REGION Network 19: EM - Execute State Complete
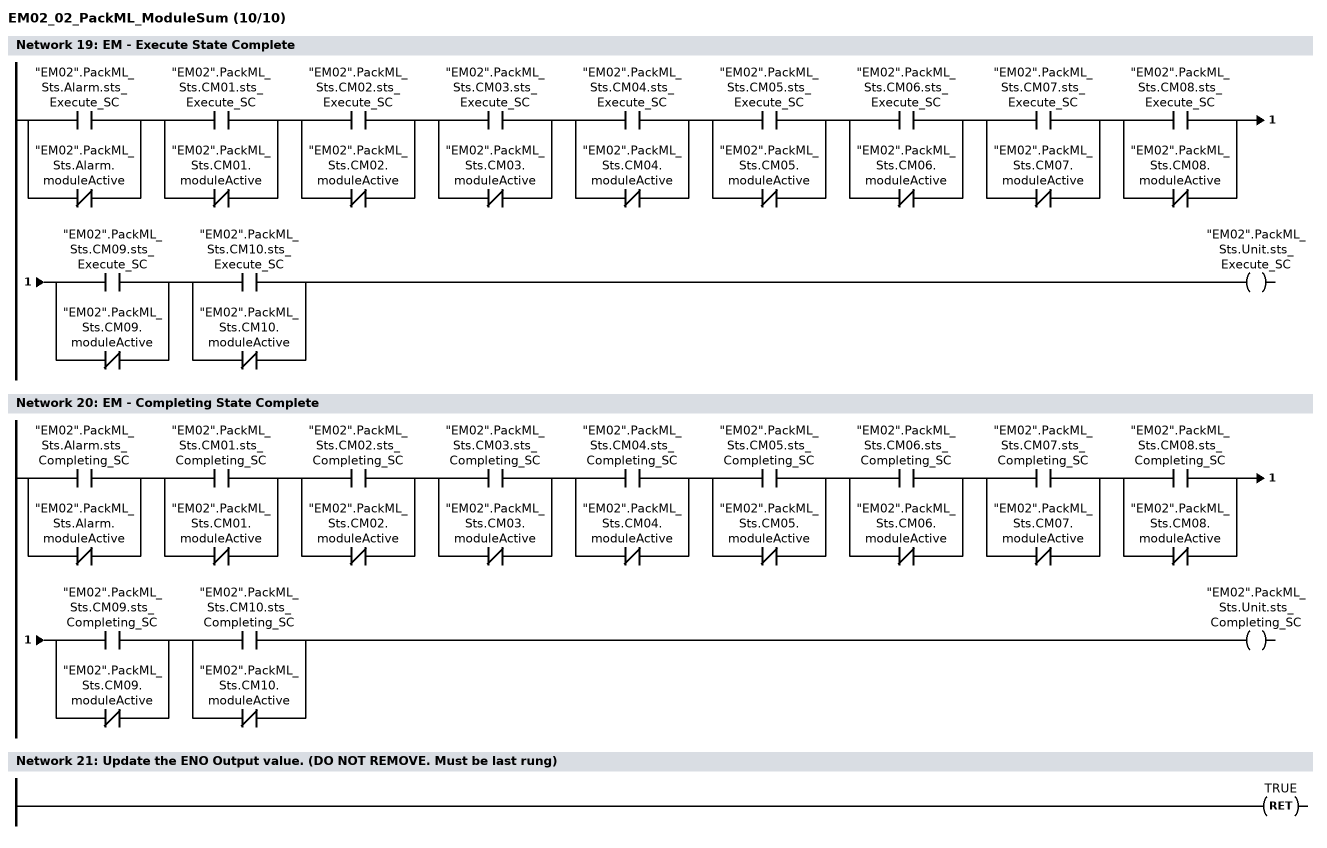
   RUNG wire#powerrail
      Contact( "EM02".PackML_Sts.Alarm.sts_Execute_SC )
      wire#w1
      Contact( "EM02".PackML_Sts.CM01.sts_Execute_SC )
      wire#w2
      Contact( "EM02".PackML_Sts.CM02.sts_Execute_SC )
      wire#w3
      Contact( "EM02".PackML_Sts.CM03.sts_Execute_SC )
      wire#w4
      Contact( "EM02".PackML_Sts.CM04.sts_Execute_SC )
      wire#w5
      Contact( "EM02".PackML_Sts.CM05.sts_Execute_SC )
      wire#w6
      Contact( "EM02".PackML_Sts.CM06.sts_Execute_SC )
      wire#w7
      Contact( "EM02".PackML_Sts.CM07.sts_Execute_SC )
      wire#w8
      Contact( "EM02".PackML_Sts.CM08.sts_Execute_SC )
      wire#w9
      Contact( "EM02".PackML_Sts.CM09.sts_Execute_SC )
      wire#w10
      Contact( "EM02".PackML_Sts.CM10.sts_Execute_SC )
      wire#w11
      Coil( "EM02".PackML_Sts.Unit.sts_Execute_SC )
   END_RUNG
   RUNG wire#powerrail
      I_Contact( "EM02".PackML_Sts.Alarm.moduleActive )
   END_RUNG wire#w1
   RUNG wire#w1
      I_Contact( "EM02".PackML_Sts.CM01.moduleActive )
   END_RUNG wire#w2
   RUNG wire#w2
      I_Contact( "EM02".PackML_Sts.CM02.moduleActive )
   END_RUNG wire#w3
   RUNG wire#w3
      I_Contact( "EM02".PackML_Sts.CM03.moduleActive )
   END_RUNG wire#w4
   RUNG wire#w4
      I_Contact( "EM02".PackML_Sts.CM04.moduleActive )
   END_RUNG wire#w5
   RUNG wire#w5
      I_Contact( "EM02".PackML_Sts.CM05.moduleActive )
   END_RUNG wire#w6
   RUNG wire#w6
      I_Contact( "EM02".PackML_Sts.CM06.moduleActive )
   END_RUNG wire#w7
   RUNG wire#w7
      I_Contact( "EM02".PackML_Sts.CM07.moduleActive )
   END_RUNG wire#w8
   RUNG wire#w8
      I_Contact( "EM02".PackML_Sts.CM08.moduleActive )
   END_RUNG wire#w9
   RUNG wire#w9
      I_Contact( "EM02".PackML_Sts.CM09.moduleActive )
   END_RUNG wire#w10
   RUNG wire#w10
      I_Contact( "EM02".PackML_Sts.CM10.moduleActive )
   END_RUNG wire#w11
   // the same network as SCL:
   "EM02".PackML_Sts.Unit.sts_Execute_SC := ("EM02".PackML_Sts.Alarm.sts_Execute_SC OR NOT "EM02".PackML_Sts.Alarm.moduleActive) AND ("EM02".PackML_Sts.CM01.sts_Execute_SC OR NOT "EM02".PackML_Sts.CM01.moduleActive) AND ("EM02".PackML_Sts.CM02.sts_Execute_SC OR NOT "EM02".PackML_Sts.CM02.moduleActive) AND ("EM02".PackML_Sts.CM03.sts_Execute_SC OR NOT "EM02".PackML_Sts.CM03.moduleActive) AND ("EM02".PackML_Sts.CM04.sts_Execute_SC OR NOT "EM02".PackML_Sts.CM04.moduleActive) AND ("EM02".PackML_Sts.CM05.sts_Execute_SC OR NOT "EM02".PackML_Sts.CM05.moduleActive) AND ("EM02".PackML_Sts.CM06.sts_Execute_SC OR NOT "EM02".PackML_Sts.CM06.moduleActive) AND ("EM02".PackML_Sts.CM07.sts_Execute_SC OR NOT "EM02".PackML_Sts.CM07.moduleActive) AND ("EM02".PackML_Sts.CM08.sts_Execute_SC OR NOT "EM02".PackML_Sts.CM08.moduleActive) AND ("EM02".PackML_Sts.CM09.sts_Execute_SC OR NOT "EM02".PackML_Sts.CM09.moduleActive) AND ("EM02".PackML_Sts.CM10.sts_Execute_SC OR NOT "EM02".PackML_Sts.CM10.moduleActive);
END_REGION

REGION Network 20: EM - Completing State Complete
   RUNG wire#powerrail
      Contact( "EM02".PackML_Sts.Alarm.sts_Completing_SC )
      wire#w1
      Contact( "EM02".PackML_Sts.CM01.sts_Completing_SC )
      wire#w2
      Contact( "EM02".PackML_Sts.CM02.sts_Completing_SC )
      wire#w3
      Contact( "EM02".PackML_Sts.CM03.sts_Completing_SC )
      wire#w4
      Contact( "EM02".PackML_Sts.CM04.sts_Completing_SC )
      wire#w5
      Contact( "EM02".PackML_Sts.CM05.sts_Completing_SC )
      wire#w6
      Contact( "EM02".PackML_Sts.CM06.sts_Completing_SC )
      wire#w7
      Contact( "EM02".PackML_Sts.CM07.sts_Completing_SC )
      wire#w8
      Contact( "EM02".PackML_Sts.CM08.sts_Completing_SC )
      wire#w9
      Contact( "EM02".PackML_Sts.CM09.sts_Completing_SC )
      wire#w10
      Contact( "EM02".PackML_Sts.CM10.sts_Completing_SC )
      wire#w11
      Coil( "EM02".PackML_Sts.Unit.sts_Completing_SC )
   END_RUNG
   RUNG wire#powerrail
      I_Contact( "EM02".PackML_Sts.Alarm.moduleActive )
   END_RUNG wire#w1
   RUNG wire#w1
      I_Contact( "EM02".PackML_Sts.CM01.moduleActive )
   END_RUNG wire#w2
   RUNG wire#w2
      I_Contact( "EM02".PackML_Sts.CM02.moduleActive )
   END_RUNG wire#w3
   RUNG wire#w3
      I_Contact( "EM02".PackML_Sts.CM03.moduleActive )
   END_RUNG wire#w4
   RUNG wire#w4
      I_Contact( "EM02".PackML_Sts.CM04.moduleActive )
   END_RUNG wire#w5
   RUNG wire#w5
      I_Contact( "EM02".PackML_Sts.CM05.moduleActive )
   END_RUNG wire#w6
   RUNG wire#w6
      I_Contact( "EM02".PackML_Sts.CM06.moduleActive )
   END_RUNG wire#w7
   RUNG wire#w7
      I_Contact( "EM02".PackML_Sts.CM07.moduleActive )
   END_RUNG wire#w8
   RUNG wire#w8
      I_Contact( "EM02".PackML_Sts.CM08.moduleActive )
   END_RUNG wire#w9
   RUNG wire#w9
      I_Contact( "EM02".PackML_Sts.CM09.moduleActive )
   END_RUNG wire#w10
   RUNG wire#w10
      I_Contact( "EM02".PackML_Sts.CM10.moduleActive )
   END_RUNG wire#w11
   // the same network as SCL:
   "EM02".PackML_Sts.Unit.sts_Completing_SC := ("EM02".PackML_Sts.Alarm.sts_Completing_SC OR NOT "EM02".PackML_Sts.Alarm.moduleActive) AND ("EM02".PackML_Sts.CM01.sts_Completing_SC OR NOT "EM02".PackML_Sts.CM01.moduleActive) AND ("EM02".PackML_Sts.CM02.sts_Completing_SC OR NOT "EM02".PackML_Sts.CM02.moduleActive) AND ("EM02".PackML_Sts.CM03.sts_Completing_SC OR NOT "EM02".PackML_Sts.CM03.moduleActive) AND ("EM02".PackML_Sts.CM04.sts_Completing_SC OR NOT "EM02".PackML_Sts.CM04.moduleActive) AND ("EM02".PackML_Sts.CM05.sts_Completing_SC OR NOT "EM02".PackML_Sts.CM05.moduleActive) AND ("EM02".PackML_Sts.CM06.sts_Completing_SC OR NOT "EM02".PackML_Sts.CM06.moduleActive) AND ("EM02".PackML_Sts.CM07.sts_Completing_SC OR NOT "EM02".PackML_Sts.CM07.moduleActive) AND ("EM02".PackML_Sts.CM08.sts_Completing_SC OR NOT "EM02".PackML_Sts.CM08.moduleActive) AND ("EM02".PackML_Sts.CM09.sts_Completing_SC OR NOT "EM02".PackML_Sts.CM09.moduleActive) AND ("EM02".PackML_Sts.CM10.sts_Completing_SC OR NOT "EM02".PackML_Sts.CM10.moduleActive);
END_REGION

REGION Network 21: Update the ENO Output value. (DO NOT REMOVE. Must be last rung)
   RUNG wire#powerrail
      ReturnCoil( TRUE )
   END_RUNG
   // the same network as SCL:
   ENO := TRUE;
   RETURN;
END_REGION
END_FUNCTION_BLOCK

FUNCTION_BLOCK "EM02_CM01_Conveyor"   // FB31691, LAD
TITLE = EM02_CM01
{ S7_Optimized_Access := 'TRUE' }
AUTHOR : tech.team.motioncontrol@siemens.com
FAMILY : CPG
VERSION : 1.1
// Support: tech.team.motioncontrol@siemens.com
   VAR
      statDummyBool : Bool;   // dummy bool - placeholder
      instBeltConveyor : "BeltConveyor";
   END_VAR
BEGIN

REGION Network 1: *** Begin the Setpoint Management Information Section ***
END_REGION

REGION Network 2: *** Begin the Logic Section ***
END_REGION

REGION Network 3: EM02_CM01_Conveyor
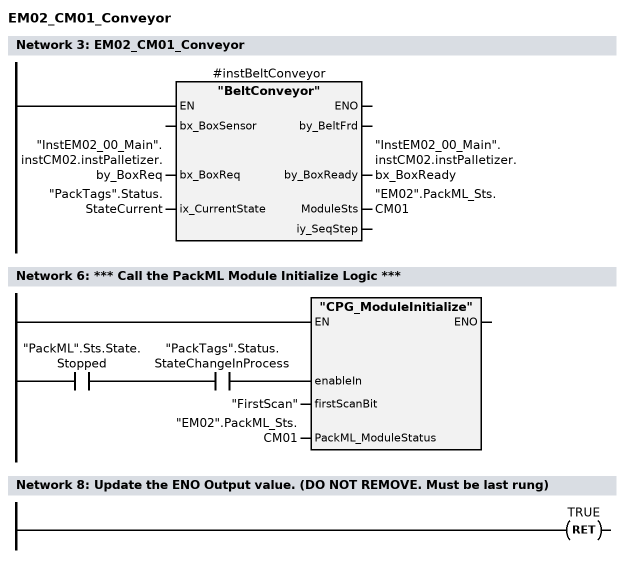
   RUNG wire#powerrail
      #instBeltConveyor(bx_BoxSensor :=, bx_BoxReq := "InstEM02_00_Main".instCM02.instPalletizer.by_BoxReq, ix_CurrentState := "PackTags".Status.StateCurrent, by_BeltFrd =>, by_BoxReady => "InstEM02_00_Main".instCM02.instPalletizer.bx_BoxReady, ModuleSts => "EM02".PackML_Sts.CM01, iy_SeqStep =>)
   END_RUNG
   // the same network as SCL:
   #instBeltConveyor(bx_BoxReq := "InstEM02_00_Main".instCM02.instPalletizer.by_BoxReq,   // "BeltConveyor"
                     ix_CurrentState := "PackTags".Status.StateCurrent,
                     by_BoxReady => "InstEM02_00_Main".instCM02.instPalletizer.bx_BoxReady,
                     ModuleSts => "EM02".PackML_Sts.CM01);
END_REGION

REGION Network 4: *** Begin the Event Information Section ***
END_REGION

REGION Network 5: *** Begin the State Model Status Feedback Section ***
END_REGION

REGION Network 6: *** Call the PackML Module Initialize Logic ***
   RUNG wire#powerrail
      "CPG_ModuleInitialize"(enableIn := wire#w1, firstScanBit := "FirstScan", PackML_ModuleStatus := "EM02".PackML_Sts.CM01)
   END_RUNG
   RUNG wire#powerrail
      Contact( "PackML".Sts.State.Stopped )
      Contact( "PackTags".Status.StateChangeInProcess )
   END_RUNG wire#w1
   // the same network as SCL:
   "CPG_ModuleInitialize"(enableIn := "PackML".Sts.State.Stopped AND "PackTags".Status.StateChangeInProcess,
                          firstScanBit := "FirstScan",
                          PackML_ModuleStatus := "EM02".PackML_Sts.CM01);
END_REGION

REGION Network 8: Update the ENO Output value. (DO NOT REMOVE. Must be last rung)
   RUNG wire#powerrail
      ReturnCoil( TRUE )
   END_RUNG
   // the same network as SCL:
   ENO := TRUE;
   RETURN;
END_REGION
END_FUNCTION_BLOCK

FUNCTION_BLOCK "EM02_CM02_Palletizer"   // FB31692, LAD
TITLE = EM02_CM02
{ S7_Optimized_Access := 'TRUE' }
AUTHOR : tech.team.motioncontrol@siemens.com
FAMILY : CPG
VERSION : 1.1
// Support: tech.team.motioncontrol@siemens.com
   VAR
      statDummyBool : Bool;   // dummy bool - placeholder
      instPalletizer : "Palletizer";
      boxCounterNTrig : Bool;
   END_VAR
BEGIN

REGION Network 1: *** Begin the Setpoint Management Information Section ***
END_REGION

REGION Network 2: *** Begin the Logic Section ***
END_REGION

REGION Network 3: *** Begin the Event Information Section ***
END_REGION

REGION Network 4: *** Begin the State Model Status Feedback Section ***
END_REGION

REGION Network 5: *** Call the PackML Module Initialize Logic ***
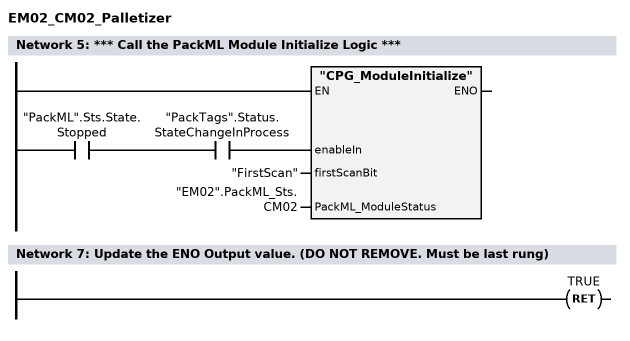
   RUNG wire#powerrail
      "CPG_ModuleInitialize"(enableIn := wire#w1, firstScanBit := "FirstScan", PackML_ModuleStatus := "EM02".PackML_Sts.CM02)
   END_RUNG
   RUNG wire#powerrail
      Contact( "PackML".Sts.State.Stopped )
      Contact( "PackTags".Status.StateChangeInProcess )
   END_RUNG wire#w1
   // the same network as SCL:
   "CPG_ModuleInitialize"(enableIn := "PackML".Sts.State.Stopped AND "PackTags".Status.StateChangeInProcess,
                          firstScanBit := "FirstScan",
                          PackML_ModuleStatus := "EM02".PackML_Sts.CM02);
END_REGION

REGION Network 7: Update the ENO Output value. (DO NOT REMOVE. Must be last rung)
   RUNG wire#powerrail
      ReturnCoil( TRUE )
   END_RUNG
   // the same network as SCL:
   ENO := TRUE;
   RETURN;
END_REGION
END_FUNCTION_BLOCK

// folder: OrganizationBlocks (OBs)

ORGANIZATION_BLOCK "CYC_INT5"   // OB35, LAD, CyclicInterrupt
TITLE = "Cyclic Interrupt"
{ S7_Optimized_Access := 'TRUE' }
VERSION : 0.1
   VAR_INPUT
      Initial_Call : Bool;   // Initial call of this OB
      Event_Count : Int;   // Events discarded
   END_VAR
BEGIN
END_ORGANIZATION_BLOCK

ORGANIZATION_BLOCK "Time error interrupt"   // OB80, LAD, TimeErrorInterrupt
{ S7_Optimized_Access := 'TRUE' }
VERSION : 0.1
   VAR_INPUT
      Fault_ID : Byte;   // Fault identifier
      Csg_OBnr : OB_Any;   // Number of OB causing the error
      Csg_Prio : UInt;   // Priority of OB causing the error
   END_VAR
BEGIN
END_ORGANIZATION_BLOCK

ORGANIZATION_BLOCK "I/O_FLT1"   // OB82, LAD, DiagnosticErrorInterrupt
TITLE = "I/O Point Fault"
{ S7_Optimized_Access := 'TRUE' }
VERSION : 0.1
   VAR_INPUT
      IO_State : Word;   // IO state of the HW object
      LADDR : Hw_Any;   // Hardware identifier
      Channel : UInt;   // Channel number
      MultiError : Bool;   // =true if more than one error is present
   END_VAR
BEGIN
END_ORGANIZATION_BLOCK

ORGANIZATION_BLOCK "I/O_FLT2"   // OB83, LAD, PullPlug
TITLE = "I/O Point Fault"
{ S7_Optimized_Access := 'TRUE' }
VERSION : 0.1
   VAR_INPUT
      LADDR : Hw_Io;   // Hardware identifier
      Event_Class : Byte;   // 16#38/39: module inserted, removed
      Fault_ID : Byte;   // Fault identifier
   END_VAR
BEGIN
END_ORGANIZATION_BLOCK

ORGANIZATION_BLOCK "RACK_FLT"   // OB86, LAD, RackStationFailure
TITLE = "Loss Of Rack Fault"
{ S7_Optimized_Access := 'TRUE' }
VERSION : 0.1
   VAR_INPUT
      LADDR : Hw_Io;   // Hardware identifier
      Event_Class : Byte;   // Event class
      Fault_ID : Byte;   // Fault identifier
   END_VAR
   VAR_TEMP
      OB86_RACKS_FLTD : Array[0..31] of Bool;
      OB86_DATE_TIME : Date_And_Time;   // Date and time OB86 started
   END_VAR
BEGIN
END_ORGANIZATION_BLOCK

ORGANIZATION_BLOCK "COMPLETE RESTART"   // OB100, LAD, Startup
TITLE = "Complete Restart"
{ S7_Optimized_Access := 'TRUE' }
VERSION : 0.1
   VAR_INPUT
      LostRetentive : Bool;   // True if retentive data are lost
      LostRTC : Bool;   // True if date and time are lost
   END_VAR
BEGIN
END_ORGANIZATION_BLOCK

ORGANIZATION_BLOCK "Programming error"   // OB121, LAD, ProgrammingError
{ S7_Optimized_Access := 'TRUE' }
VERSION : 0.1
   VAR_INPUT
      BlockNr : UInt;   // Number of causing block
      Reaction : USInt;   // 0:ignore, 1:substitute, 2:skip
      Fault_ID : Byte;   // Fault identifier
      BlockType : USInt;   // 16#01:OB, 16#02:FC, 16#03:FB, 16#04:SFC, 16#05:SFB, 16#06:DB: Type of block causing the error
      Area : USInt;   // Area where the error occured
      DBNr : DB_ANY;   // DB number if Area = DB or DI
      Csg_OBNr : OB_Any;   // Number of OB causing the error
      Csg_Prio : USInt;   // Priority of OB causing the error
      Width : USInt;   // 0:bit, 1:byte, 2:word, 3:dword, 4:lword
   END_VAR
BEGIN
END_ORGANIZATION_BLOCK

// folder: SupportingBlocks/CPG_Blocks

FUNCTION_BLOCK "CPG_AlarmHistory"   // FB31600, SCL
TITLE = CPG_AlarmHistory
{ S7_Optimized_Access := 'TRUE' }
AUTHOR : tech.team.motioncontrol@siemens.com
FAMILY : CPG
VERSION : 1.1
// Support: tech.team.motioncontrol@siemens.com
   VAR_OUTPUT
      alarmHistoryArraySize : Int;   // Size of Alarm History - number of alarm array elements
   END_VAR
   VAR_IN_OUT
      inStopReasonAlarm : "CPG_typeEvent";   // Input - Stop Reason Alarm (structure)
      stsAlarmHistory : Array[0.."CPG_NO_OF_ADMIN_EVENTS_HISTORY_UPPER_LIM"] of "CPG_typeEvent";   // Status- Alarm History Log
   END_VAR
   VAR
      statAlarmArraySize : Int;   // Max # of Events in the Alarm History Array
      statTriggerOsPos : Bool;   // Trigger One Shot - positive edge
      statTriggerOsNeg : Bool;   // Trigger One Shot - negative edge
      statErrorRtc : Int;   // Error code for reading of Real Time Clock
      statEventCurDateTime : DTL;   // temp value for current date & time
      statFirstScan : Bool;   // 0=1st scan of FB; set to 1 after 1st FB scan...
   END_VAR
   VAR_TEMP
      tempIndex : Int;   // temp index value
   END_VAR
   VAR CONSTANT
      ZERO : Int := 0;   // constant = 0
      NEGATIVE_ONE : Int := -1;   // constant = -1
   END_VAR
BEGIN
   //============================================================================================================
   // SIEMENS AG
   // (c)Copyright 2018 All Rights Reserved
   //------------------------------------------------------------------------------------------------------------
   // Project: CPG Template
   // Tested with: S7-1500 with FW version V2.1
   // Engineering: TIA Portal V14
   // Restrictions: ---
   // Requirements: S7-1500
   // Functionality: used to capture the current Stop ReasonAlarm (i.e. 'Machine)
   //                First Fault to the "PackTags" AlarmHistory log.
   // Support: tech.team.motioncontrol@siemens.com
   //------------------------------------------------------------------------------------------------------------
   // Change log table:
   // Version       Date               Expert in charge    Changes applied
   //  01.00.00     01.01.2018         MP                  Initial Release & PackML V1.5  Renamed CPG V1.0
   //  01.01.00     22.05.2018         JP                  Adopted to styleguide
   //  01.01.01     01.05.2020         KB                  Changed RD_SYS_T -> RD_LOC_T
   //============================================================================================================
   // Function : CPG_AlarmHistory
   //============================================================================================================

   // First Scan Logic
   IF #statFirstScan = FALSE THEN
     "CPG_ArrayLength"(arrayToBeSized := #stsAlarmHistory,
                       arraySize => #statAlarmArraySize);

     // Update number of array elements in Alarm History Array (used for Admin.AlarmHistoryExtent)
     #alarmHistoryArraySize := #statAlarmArraySize;

     #statFirstScan := TRUE;      // Set the FB 1st Scan Bit
   END_IF;

   // Positive Trigger
   IF #inStopReasonAlarm.Trigger = TRUE AND #statTriggerOsPos = FALSE THEN
     // execute code for new incoming event
     #statTriggerOsPos := TRUE;   // Set the One Shot Bit 

     // Index the existing Alarm History Array (FIFO).
     FOR #tempIndex := #statAlarmArraySize - 1 TO 1 BY -1 DO
       #stsAlarmHistory[#tempIndex] := #stsAlarmHistory[#tempIndex - 1];
     END_FOR;

     // Update the Array[0] with the current alarm information
     #stsAlarmHistory[0] := #inStopReasonAlarm;
   END_IF;

   IF #inStopReasonAlarm.Trigger = FALSE AND #statTriggerOsPos = TRUE THEN
     // Reset the One Shot Bit
     #statTriggerOsPos := FALSE;  // Reset the One Shot Bit
   END_IF;

   // Negative Trigger
   IF #inStopReasonAlarm.Trigger = FALSE AND #statTriggerOsNeg = FALSE THEN
     // Execute code for new incoming event
     #statTriggerOsNeg := TRUE;    // Set the One Shot Bit
     // Capture the Alarm Ack. Time
     #statErrorRtc := RD_LOC_T(#statEventCurDateTime);     // Read the Real Time Clock
     #stsAlarmHistory[0].AckDateTimeDTL := #statEventCurDateTime; // Update acknowledge time
   END_IF;

   IF #inStopReasonAlarm.Trigger = TRUE AND #statTriggerOsPos = TRUE THEN
     // Reset the One Shot Bit
     #statTriggerOsNeg := FALSE;   // Reset the One Shot Bit
   END_IF;

   //  -------------- END OF LOGIC -------------------------
   ENO := TRUE;   // Set the ENO output
END_FUNCTION_BLOCK

FUNCTION_BLOCK "CPG_AlarmMove"   // FB31601, SCL
TITLE = CPG_AlarmMove
{ S7_Optimized_Access := 'TRUE' }
AUTHOR : tech.team.motioncontrol@siemens.com
FAMILY : CPG
VERSION : 1.0
// Support: tech.team.motioncontrol@siemens.com
   VAR_INPUT
      Sts_NumEvents : Int;   // Number of Active Alarms
   END_VAR
   VAR_OUTPUT
      Sts_Error : Bool;   // Error Status. 0=no error, 1=error
      Sts_ErrorCode : Int;   // Error code / number
   END_VAR
   VAR_IN_OUT
      source : Array[0.."CPG_NO_OF_STS_ELEMENTS_EVENT_SUM_UPPER_LIM"] of "CPG_typeEvent";   // source location of the machine alarms
      destination : Array[0.."CPG_NO_OF_ADMIN_EVENTS_UPPER_LIM"] of "CPG_typeEvent";   // destination location of the PackTag alarms
   END_VAR
   VAR
      statSourceNumEvents : Int;   // MAX # OF Events - source event list
      statDestinationNumEvents : Int;   // MAX # OF Events - destination event list
      statIndex : Int;   // index value
      statPrevNumEvents : Int;   // previous number of events
      statZeroEvent : "CPG_typeEvent";   // blank event
      statWrkNumEvents : Int;   // working number of active events
   END_VAR
BEGIN
   //============================================================================================================
   // SIEMENS AG
   // (c)Copyright 2018 All Rights Reserved
   //------------------------------------------------------------------------------------------------------------
   // Project: CPG Template
   // Tested with: S7-1500 with FW version V2.1
   // Engineering: TIA Portal V14
   // Restrictions: ---
   // Requirements: S7-1500
   // Functionality: move alarm structures 
   // Support: tech.team.motioncontrol@siemens.com
   //------------------------------------------------------------------------------------------------------------
   // Change log table:
   // Version       Date               Expert in charge    Changes applied
   //  01.00.00     01.01.2018         MP                  Initial Release & PackML V1.5  Renamed CPG V1.0
   //  01.01.00     22.05.2018         JP                  Adopted to styleguide
   //============================================================================================================
   // Function : CPG_AlarmMove
   //============================================================================================================


   // initialize & determine max array size
   "CPG_ArrayLength"(arrayToBeSized := #source,
                     arraySize => #statSourceNumEvents);

   "CPG_ArrayLength"(arrayToBeSized := #destination,
                     arraySize => #statDestinationNumEvents);

   #statWrkNumEvents := #Sts_NumEvents;

   IF (#statDestinationNumEvents < #statSourceNumEvents) AND (#statDestinationNumEvents < #Sts_NumEvents) THEN
     #statWrkNumEvents := #statDestinationNumEvents;
   END_IF;

   IF (#statSourceNumEvents < #statDestinationNumEvents) AND (#statSourceNumEvents < #Sts_NumEvents) THEN
     #statWrkNumEvents := #statSourceNumEvents;
   END_IF;

   FOR #statIndex := 0 TO #statWrkNumEvents - 1 DO
     #destination[#statIndex] := #source[#statIndex];
   END_FOR;

   // Clean up event list
   IF #statPrevNumEvents > #statWrkNumEvents THEN
     FOR #statIndex := #statWrkNumEvents TO #statPrevNumEvents - 1 DO
       #destination[#statIndex] := #statZeroEvent;
     END_FOR;
   END_IF;

   #statPrevNumEvents := #statWrkNumEvents;

   //  -------------- END OF LOGIC -------------------------
   ENO := TRUE;   // Set the ENO output
END_FUNCTION_BLOCK

FUNCTION_BLOCK "CPG_Event"   // FB31602, SCL
TITLE = CPG_Event
{ S7_Optimized_Access := 'TRUE' }
AUTHOR : tech.team.motioncontrol@siemens.com
FAMILY : CPG
VERSION : 1.1
// Support: tech.team.motioncontrol@siemens.com
   VAR_INPUT
      EnableIn : Bool;   // Enable the FB call.
      Cfg_Event : "CPG_typeEventCfg";   // configuration data structure for this event
      Cfg_MessagePrefix : "CPG_typeMessagePrefix";   // Message Prefix value for event messages
   END_VAR
   VAR_OUTPUT
      Sts_Active : Bool;   // event is currently active
      Sts_Latched : Bool;   // event has been active since last reset command
   END_VAR
   VAR_IN_OUT
      In_EventStatus : "CPG_typeEventStatus";   // Working event list data section
   END_VAR
   VAR
      statActive : Bool;   // event is currently active
      statLatched : Bool;   // event has been active since last reset command
      statEvent_Number : Int;   // Event Number
      statPrev_ResetID : Int;   // Prev Reset ID
      statError_RTC : Int;   // Error code for reading of Real Time Clock
      statEvent_CurDateTime : DTL;   // temp value for current date & time
   END_VAR
   VAR_TEMP
      tempLanguage : Int;   // value of the currently selected language
   END_VAR
BEGIN
   //============================================================================================================
   // SIEMENS AG
   // (c)Copyright 2018 All Rights Reserved
   //------------------------------------------------------------------------------------------------------------
   // Project: CPG Template
   // Tested with: S7-1500 with FW version V2.1
   // Engineering: TIA Portal V14
   // Restrictions: ---
   // Requirements: S7-1500
   // Functionality: Control TR88 EVENT functions for CPG Template. 
   // Support: tech.team.motioncontrol@siemens.com
   //------------------------------------------------------------------------------------------------------------
   // Change log table:
   // Version       Date               Expert in charge    Changes applied
   //  01.00.00     01.01.2018         MP                  Initial Release & PackML V1.8  Renamed CPG V1.0
   //  01.01.00     22.05.2018         JP                  Adopted to styleguide
   //  01.01.01     06.02.2020         KB                  Optimized call of Concat instruction
   //                                                      Changed RD_SYS_T -> RD_LOC_T
   //============================================================================================================
   // Function : CPG_Event
   //============================================================================================================

   // ===========================================================================
   //  Begin the LOGIC section:

   //-------------  If ENABLE is FALSE----------------------------------------
   IF NOT (#EnableIn) THEN                          // If block is not enabled, then
     IF #statActive THEN              // Status Active
       IF #statEvent_Number < #In_EventStatus.wrk_EventArraySize THEN   // current event below max size?
         #statError_RTC := RD_LOC_T(#statEvent_CurDateTime);            // Read the Real Time Clock
         #In_EventStatus.sts_Events[#statEvent_Number].AckDateTimeDTL := #statEvent_CurDateTime; // update Acknowledge time
         #In_EventStatus.sts_Events[#statEvent_Number].Trigger := FALSE;
       END_IF;                     // IF Event_Number

       #statActive := FALSE;             // Reset the active bit        
       #In_EventStatus.wrk_UpdateEventListID := #In_EventStatus.wrk_UpdateEventListID + 1;
     END_IF;                             // IF Sts_Active

     IF #statLatched AND (#In_EventStatus.wrk_ResetID <> #statPrev_ResetID) THEN
       #statLatched := FALSE;
       #In_EventStatus.wrk_UpdateEventListID := #In_EventStatus.wrk_UpdateEventListID + 1;
       #statPrev_ResetID := #In_EventStatus.wrk_ResetID;
     END_IF;             // IF Sts_Latched

     ENO := FALSE;         // enable out is false (0)

   ELSE                    // else IF NOT (enable)
     //-------------  If ENABLE is TRUE ----------------------------------------  
     // If this FB is enabled....  
     IF NOT (#statActive) OR (#In_EventStatus.wrk_ResetID <> #statPrev_ResetID) THEN
       IF NOT (#statLatched) THEN
         #statError_RTC := RD_LOC_T(#statEvent_CurDateTime);            // Read the Real Time Clock
       END_IF;

       IF NOT (#statLatched) OR (#In_EventStatus.wrk_ResetID <> #statPrev_ResetID) THEN
         #statEvent_Number := #In_EventStatus.sts_NumAllEvents;             // increment event number
         #In_EventStatus.sts_NumAllEvents := #In_EventStatus.sts_NumAllEvents + 1;         // increment number of all event
         #statPrev_ResetID := #In_EventStatus.wrk_ResetID;                                     // update previous Reset ID      
       END_IF;

       IF #statEvent_Number < #In_EventStatus.wrk_EventArraySize THEN
         #tempLanguage := #In_EventStatus.wrk_LanguageSelection;

         #In_EventStatus.sts_Events[#statEvent_Number].ID := #Cfg_Event.ID;
         #In_EventStatus.sts_Events[#statEvent_Number].Value := #Cfg_Event.value;
         #In_EventStatus.sts_Events[#statEvent_Number].Category := #Cfg_Event.category;

         // update the event message String with "UN"/EM prefix + CM prefix + event message for selected language
         IF #tempLanguage >= 0 AND #tempLanguage <= "LPMLV30_LANGUAGES_UPPER_LIM" THEN
             #In_EventStatus.sts_Events[#statEvent_Number].Message := CONCAT(IN1 := #In_EventStatus.wrk_MessagePrefix,
                                                                             IN2 := #Cfg_MessagePrefix.messagePrefix[#tempLanguage], IN3 := #Cfg_Event.message[#tempLanguage]);
         ELSE
             #In_EventStatus.sts_Events[#statEvent_Number].Message := #In_EventStatus.wrk_MessagePrefix;
         END_IF;


         #In_EventStatus.sts_Events[#statEvent_Number].Trigger := TRUE;                          // Set trigger to 1 
         #In_EventStatus.sts_Events[#statEvent_Number].DateTimeDTL := #statEvent_CurDateTime;       // Update with the current time
         #In_EventStatus.sts_Events[#statEvent_Number].AckDateTimeDTL := DT#1990-1-1-0:0:0.0;       // clear the acknowledge time value 
       END_IF;

       #statActive := TRUE;                            // set the status active bit
       #statLatched := TRUE;                            // set the status latched bit
       #In_EventStatus.wrk_UpdateEventListID := #In_EventStatus.wrk_UpdateEventListID + 1;  // increment the work update listID

       CASE DINT_TO_INT(#Cfg_Event.category) OF                     // set the appropriate category lateched bit
         0:
           #In_EventStatus.sts_Category_0_Latched := TRUE;
         1:
           #In_EventStatus.sts_Category_1_Latched := TRUE;
         2:
           #In_EventStatus.sts_Category_2_Latched := TRUE;
         3:
           #In_EventStatus.sts_Category_3_Latched := TRUE;
         4:
           #In_EventStatus.sts_Category_4_Latched := TRUE;
         5:
           #In_EventStatus.sts_Category_5_Latched := TRUE;
         6:
           #In_EventStatus.sts_Category_6_Latched := TRUE;
         7:
           #In_EventStatus.sts_Category_7_Latched := TRUE;
         8:
           #In_EventStatus.sts_Category_8_Latched := TRUE;
         9:
           #In_EventStatus.sts_Category_9_Latched := TRUE;
       END_CASE;
     END_IF; // End "IF NOT (Sts_Active)"

   END_IF; // End "IF NOT(EnableIn) "

   // Write output variables
   #Sts_Latched := #statLatched;
   #Sts_Active := #statActive;

   //  -------------- END OF LOGIC -------------------------
   ENO := TRUE;   // Set the ENO output
END_FUNCTION_BLOCK

FUNCTION_BLOCK "CPG_EventManager"   // FB31603, SCL
TITLE = CPG_EventManager
{ S7_Optimized_Access := 'TRUE' }
AUTHOR : tech.team.motioncontrol@siemens.com
FAMILY : CPG
VERSION : 1.0
// Support: tech.team.motioncontrol@siemens.com
   VAR_INPUT
      Cmd_Reset : Bool;   // Reset Command
      Cmd_ClearFirstOutEvents : Bool;   // Command to clear First Out events
      firstScanBit : Bool;   // Bit used to tell logic that this is the first scan of PLC
      Cfg_MessagePrefix : "CPG_typeMessagePrefix";   // Message Prefix value for event messages multi-lingual
      Cfg_LanguageSelection : Int;   // Current Langage: 0=EN, 1=DE, 2=SP/ES, 3=IT, 4=FR
   END_VAR
   VAR_OUTPUT
      Sts_Category_0_Latched : Bool;   // Event Category Status (on until reset cmd) - CAT 0
      Sts_Category_1_Latched : Bool;   // Event Category Status (on until reset cmd) - CAT 1
      Sts_Category_2_Latched : Bool;   // Event Category Status (on until reset cmd) - CAT 2
      Sts_Category_3_Latched : Bool;   // Event Category Status (on until reset cmd) - CAT 3
      Sts_Category_4_Latched : Bool;   // Event Category Status (on until reset cmd) - CAT 4
      Sts_Category_5_Latched : Bool;   // Event Category Status (on until reset cmd) - CAT 5
      Sts_Category_6_Latched : Bool;   // Event Category Status (on until reset cmd) - CAT 6
      Sts_Category_7_Latched : Bool;   // Event Category Status (on until reset cmd) - CAT 7
      Sts_Category_8_Latched : Bool;   // Event Category Status (on until reset cmd) - CAT 8
      Sts_Category_9_Latched : Bool;   // Event Category Status (on until reset cmd) - CAT 9
      Sts_Category_0_NotLatched : Bool;   // Event Cat Status, not latched (=active event status) - CAT 0
      Sts_Category_1_NotLatched : Bool;   // Event Cat Status, not latched (=active event status) - CAT 1
      Sts_Category_2_NotLatched : Bool;   // Event Cat Status, not latched (=active event status) - CAT 2
      Sts_Category_3_NotLatched : Bool;   // Event Cat Status, not latched (=active event status) - CAT 3
      Sts_Category_4_NotLatched : Bool;   // Event Cat Status, not latched (=active event status) - CAT 4
      Sts_Category_5_NotLatched : Bool;   // Event Cat Status, not latched (=active event status) - CAT 5
      Sts_Category_6_NotLatched : Bool;   // Event Cat Status, not latched (=active event status) - CAT 6
      Sts_Category_7_NotLatched : Bool;   // Event Cat Status, not latched (=active event status) - CAT 7
      Sts_Category_8_NotLatched : Bool;   // Event Cat Status, not latched (=active event status) - CAT 8
      Sts_Category_9_NotLatched : Bool;   // Event Cat Status, not latched (=active event status) - CAT 9
      Sts_NumEvents : Int;   // Number of event in the In_EventStatus list
      Sts_CurrentActiveEvent : Bool;   // Status - TRUE = if any active events
      Sts_Error : Bool;   // FB Error exist
      Sts_ErrorCode : DInt;   // FB Error code
   END_VAR
   VAR_IN_OUT
      In_EventStatus : "CPG_typeEventStatus";   // Working event list data section
   END_VAR
   VAR
      statEventCategory : DInt;
      statIndexAllEvents : Int;
      statIndexClearActiveEvents : Int;
      statIndexClearFirstOut : Int;
      statNumEvents : Int;   // Max # of Events
      statPrevCmdReset : Bool;
      statPrevNumEvents : Int;
      statPrevUpdateEventListID : Int;
      statUpdateEventList : Bool;
      statCurrentErrorCode : Int;
      statCurrentActiveEvent : Bool;
      statZeroEvent : "CPG_typeEvent";   // Null Event
   END_VAR
BEGIN
   //============================================================================================================
   // SIEMENS AG
   // (c)Copyright 2018 All Rights Reserved
   //------------------------------------------------------------------------------------------------------------
   // Project: CPG Template
   // Tested with: S7-1500 with FW version V2.1
   // Engineering: TIA Portal V14
   // Restrictions: ---
   // Requirements: S7-1500
   // Functionality: Control EventManager function
   // Support: tech.team.motioncontrol@siemens.com
   //------------------------------------------------------------------------------------------------------------
   // Change log table:
   // Version       Date               Expert in charge    Changes applied
   //  01.00.00     01.01.2018         MP                  Initial Release & PackML V1.8  Renamed CPG V1.0
   //  01.01.00     22.05.2018         JP                  Adopted to styleguide
   //============================================================================================================
   // Function : CPG_EventManager
   //============================================================================================================

   // First Scan Logic Logic (only run through on 1st scan of PLC)
   IF #firstScanBit THEN                                                                   // Only run first scan
     #In_EventStatus.wrk_ResetID := #In_EventStatus.wrk_ResetID + 1;                     // increment the Work Reset ID
     #In_EventStatus.wrk_UpdateEventListID := #In_EventStatus.wrk_UpdateEventListID + 1; // increment the Work UpdateList ID
     #In_EventStatus.sts_NumAllEvents := 0;                                              // Reset the number of all events value

     // Determine the Number of Sts_Events for given alarm/warning area
     "CPG_ArrayLength"(arrayToBeSized := #In_EventStatus.sts_Events,
                       arraySize => #In_EventStatus.wrk_EventArraySize);
     RETURN;     // Exit the FB call
   END_IF;         // End the first scan section


   //---------------------------------------------------------------------------------
   // Main Logic Section

   // Update the message prefix for the current language
   IF #Cfg_LanguageSelection >= 0 AND #Cfg_LanguageSelection <= "LPMLV30_LANGUAGES_UPPER_LIM" THEN
     #In_EventStatus.wrk_MessagePrefix := #Cfg_MessagePrefix.messagePrefix[#Cfg_LanguageSelection];
   END_IF;
   #In_EventStatus.wrk_LanguageSelection := #Cfg_LanguageSelection;

   // Upon a reset command, reset the latched status bits and clear the event list
   IF #Cmd_Reset THEN
     #In_EventStatus.sts_Category_0_Latched := FALSE;
     #In_EventStatus.sts_Category_1_Latched := FALSE;
     #In_EventStatus.sts_Category_2_Latched := FALSE;
     #In_EventStatus.sts_Category_3_Latched := FALSE;
     #In_EventStatus.sts_Category_4_Latched := FALSE;
     #In_EventStatus.sts_Category_5_Latched := FALSE;
     #In_EventStatus.sts_Category_6_Latched := FALSE;
     #In_EventStatus.sts_Category_7_Latched := FALSE;
     #In_EventStatus.sts_Category_8_Latched := FALSE;
     #In_EventStatus.sts_Category_9_Latched := FALSE;

     IF NOT (#statPrevCmdReset) THEN                             // Clear the zero event
       #In_EventStatus.out_ZeroEvent := #statZeroEvent;
       // String seperation variable not added.
     END_IF;
   END_IF;                      // End IF Cmd_Reset.... 


   // Clear first out events - for alarms, this is typically done once the machine starts    
   IF #Cmd_ClearFirstOutEvents AND NOT (#statCurrentActiveEvent) THEN
     #In_EventStatus.sts_FirstOutEvent := #In_EventStatus.out_ZeroEvent;

     FOR #statIndexClearFirstOut := 0 TO 9 BY 1 DO
       #In_EventStatus.sts_FirstOutEventCat[#statIndexClearFirstOut] := #In_EventStatus.out_ZeroEvent;
     END_FOR;
   END_IF;

   // Determine the maximum number of event that can be stored in the array.
   // It is assumed that the input array size is equal to the output array size
   IF (#Cmd_Reset AND (NOT #statPrevCmdReset)) OR (#In_EventStatus.wrk_EventArraySize = 0) THEN
     // Determine the Number of Sts_Events for given alarm/warning area

     "CPG_ArrayLength"(arrayToBeSized := #In_EventStatus.sts_Events,
                       arraySize => #In_EventStatus.wrk_EventArraySize);
   END_IF;

   //Determine if the event list needs updating    
   IF #In_EventStatus.wrk_UpdateEventListID <> #statPrevUpdateEventListID THEN
     #statPrevUpdateEventListID := #In_EventStatus.wrk_UpdateEventListID;
     #statUpdateEventList := TRUE;
   END_IF;

   IF #statUpdateEventList THEN
     #statUpdateEventList := FALSE;
     // Update Event outputs and status
     // First clear the not latched staus bits and total number of events.
     // This instruction will find the events in the coming rungs
     #statCurrentErrorCode := 0;
     #Sts_NumEvents := #In_EventStatus.sts_NumAllEvents;
     #statCurrentActiveEvent := FALSE;
     #Sts_Category_0_NotLatched := FALSE;
     #Sts_Category_1_NotLatched := FALSE;
     #Sts_Category_2_NotLatched := FALSE;
     #Sts_Category_3_NotLatched := FALSE;
     #Sts_Category_4_NotLatched := FALSE;
     #Sts_Category_5_NotLatched := FALSE;
     #Sts_Category_6_NotLatched := FALSE;
     #Sts_Category_7_NotLatched := FALSE;
     #Sts_Category_8_NotLatched := FALSE;
     #Sts_Category_9_NotLatched := FALSE;

     //Determine if the number of events is greater than the max array size        
     //if so, then report error
     #statNumEvents := #In_EventStatus.sts_NumAllEvents;
     IF #statNumEvents > #In_EventStatus.wrk_EventArraySize THEN
       #statNumEvents := #In_EventStatus.wrk_EventArraySize;
       IF (#statCurrentErrorCode = 0) THEN                   // Update status error code
         #statCurrentErrorCode := 1;
       END_IF;
     END_IF;
     #In_EventStatus.sts_NumEvents := #statNumEvents;

     //Go through the event array to capture first fault event and perform string management        
     #statIndexAllEvents := 0;
     FOR #statIndexAllEvents := 0 TO #statNumEvents - 1 DO
       // Check to see if any event is currently still active
       IF (#In_EventStatus.sts_Events[#statIndexAllEvents].Trigger) THEN
         #statCurrentActiveEvent := TRUE;
       END_IF;

       //Store event category for logic later in code
       IF (#In_EventStatus.sts_Events[#statIndexAllEvents].Category >= 0) AND (#In_EventStatus.sts_Events[#statIndexAllEvents].Category <= 9) THEN
         #statEventCategory := #In_EventStatus.sts_Events[#statIndexAllEvents].Category;
       ELSE
         #statEventCategory := 0;
         IF (#statCurrentErrorCode = 0) THEN                   // Update status error code
           #statCurrentErrorCode := 2;
         END_IF;         // end "IF (Sts_ErrorCode=0)"
       END_IF;             // end "IF (In_EventStatus.Sts_Events[Inde..."    

       // Set the First Out Event
       IF NOT (#In_EventStatus.sts_FirstOutEvent.Trigger) THEN
         #In_EventStatus.sts_FirstOutEvent := #In_EventStatus.sts_Events[#statIndexAllEvents];
         #In_EventStatus.sts_FirstOutEvent.Trigger := TRUE;
       END_IF;

       // Set the First Out Events by category
       IF NOT (#In_EventStatus.sts_FirstOutEventCat[#statEventCategory].Trigger) THEN
         #In_EventStatus.sts_FirstOutEventCat[#statEventCategory] := #In_EventStatus.sts_Events[#statIndexAllEvents];
         #In_EventStatus.sts_FirstOutEventCat[#statEventCategory].Trigger := TRUE;
       END_IF;

       //Category Event Status            
       CASE DINT_TO_INT(#In_EventStatus.sts_Events[#statIndexAllEvents].Category) OF
         0:
           #Sts_Category_0_NotLatched := #In_EventStatus.sts_Events[#statIndexAllEvents].Trigger;
         1:
           #Sts_Category_1_NotLatched := (#Sts_Category_1_NotLatched OR #In_EventStatus.sts_Events[#statIndexAllEvents].Trigger);
         2:
           #Sts_Category_2_NotLatched := (#Sts_Category_2_NotLatched OR #In_EventStatus.sts_Events[#statIndexAllEvents].Trigger);
         3:
           #Sts_Category_3_NotLatched := (#Sts_Category_3_NotLatched OR #In_EventStatus.sts_Events[#statIndexAllEvents].Trigger);
         4:
           #Sts_Category_4_NotLatched := (#Sts_Category_4_NotLatched OR #In_EventStatus.sts_Events[#statIndexAllEvents].Trigger);
         5:
           #Sts_Category_5_NotLatched := (#Sts_Category_5_NotLatched OR #In_EventStatus.sts_Events[#statIndexAllEvents].Trigger);
         6:
           #Sts_Category_6_NotLatched := (#Sts_Category_6_NotLatched OR #In_EventStatus.sts_Events[#statIndexAllEvents].Trigger);
         7:
           #Sts_Category_7_NotLatched := (#Sts_Category_7_NotLatched OR #In_EventStatus.sts_Events[#statIndexAllEvents].Trigger);
         8:
           #Sts_Category_8_NotLatched := (#Sts_Category_8_NotLatched OR #In_EventStatus.sts_Events[#statIndexAllEvents].Trigger);
         9:
           #Sts_Category_9_NotLatched := (#Sts_Category_9_NotLatched OR #In_EventStatus.sts_Events[#statIndexAllEvents].Trigger);
       END_CASE;  // End of DINT_TO_INT(In_EventStatus.sts_events[Ind....


     END_FOR;

     // set the status bits
     #Sts_Category_0_Latched := #In_EventStatus.sts_Category_0_Latched;
     #Sts_Category_1_Latched := #In_EventStatus.sts_Category_1_Latched;
     #Sts_Category_2_Latched := #In_EventStatus.sts_Category_2_Latched;
     #Sts_Category_3_Latched := #In_EventStatus.sts_Category_3_Latched;
     #Sts_Category_4_Latched := #In_EventStatus.sts_Category_4_Latched;
     #Sts_Category_5_Latched := #In_EventStatus.sts_Category_5_Latched;
     #Sts_Category_6_Latched := #In_EventStatus.sts_Category_6_Latched;
     #Sts_Category_7_Latched := #In_EventStatus.sts_Category_7_Latched;
     #Sts_Category_8_Latched := #In_EventStatus.sts_Category_8_Latched;
     #Sts_Category_9_Latched := #In_EventStatus.sts_Category_9_Latched;

     #In_EventStatus.sts_Category_0_NotLatched := #Sts_Category_0_NotLatched;
     #In_EventStatus.sts_Category_1_NotLatched := #Sts_Category_1_NotLatched;
     #In_EventStatus.sts_Category_2_NotLatched := #Sts_Category_2_NotLatched;
     #In_EventStatus.sts_Category_3_NotLatched := #Sts_Category_3_NotLatched;
     #In_EventStatus.sts_Category_4_NotLatched := #Sts_Category_4_NotLatched;
     #In_EventStatus.sts_Category_5_NotLatched := #Sts_Category_5_NotLatched;
     #In_EventStatus.sts_Category_6_NotLatched := #Sts_Category_6_NotLatched;
     #In_EventStatus.sts_Category_7_NotLatched := #Sts_Category_7_NotLatched;
     #In_EventStatus.sts_Category_8_NotLatched := #Sts_Category_8_NotLatched;
     #In_EventStatus.sts_Category_9_NotLatched := #Sts_Category_9_NotLatched;

     #In_EventStatus.sts_CurrentActiveEvent := #statCurrentActiveEvent;
   END_IF;

   // Clear the remaining inactive bits    
   IF #statPrevNumEvents > #In_EventStatus.sts_NumEvents THEN
     FOR #statIndexClearActiveEvents := #In_EventStatus.sts_NumEvents TO #statPrevNumEvents - 1 DO
       #In_EventStatus.sts_Events[#statIndexClearActiveEvents] := #In_EventStatus.out_ZeroEvent;
     END_FOR;
   END_IF;

   // Clear the number of input events in the case where some control module events are not being actively scanned.    
   IF #Cmd_Reset AND ((#In_EventStatus.sts_CurrentActiveEvent) OR (#In_EventStatus.sts_NumEvents > 0) OR (NOT #statPrevCmdReset)) THEN
     #In_EventStatus.wrk_ResetID := #In_EventStatus.wrk_ResetID + 1;
     #In_EventStatus.wrk_UpdateEventListID := #In_EventStatus.wrk_UpdateEventListID + 1;
     #In_EventStatus.sts_NumAllEvents := 0;
   END_IF;

   #statPrevNumEvents := #In_EventStatus.sts_NumEvents;
   #statPrevCmdReset := #Cmd_Reset;

   //Write outputs
   #Sts_ErrorCode := #statCurrentErrorCode;
   #Sts_Error := (#statCurrentErrorCode <> 0);
   #Sts_CurrentActiveEvent := #statCurrentActiveEvent;

   //-----------------------------------------------------
   ENO := TRUE;   // Set the ENO output
END_FUNCTION_BLOCK

FUNCTION_BLOCK "CPG_EventSortFilter"   // FB31604, SCL
TITLE = CPG_EventSortFilter
{ S7_Optimized_Access := 'TRUE' }
AUTHOR : tech.team.motioncontrol@siemens.com
FAMILY : CPG